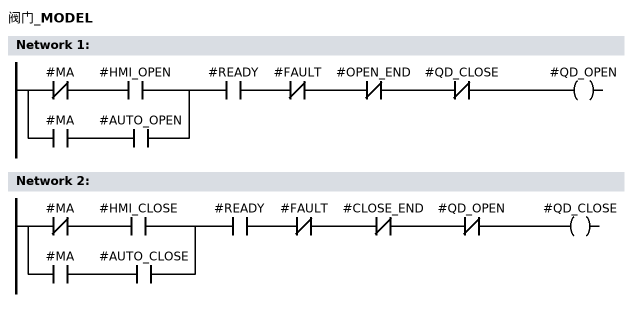
   RUNG wire#powerrail
      I_Contact( #MA )
      Contact( #HMI_OPEN )
      wire#w1
      Contact( #READY )
      I_Contact( #FAULT )
      I_Contact( #OPEN_END )
      I_Contact( #QD_CLOSE )
      Coil( #QD_OPEN )
   END_RUNG
   RUNG wire#powerrail
      Contact( #MA )
      Contact( #AUTO_OPEN )
   END_RUNG wire#w1
   // the same network as SCL:
   #QD_OPEN := ((NOT #MA AND #HMI_OPEN) OR (#MA AND #AUTO_OPEN)) AND #READY AND NOT #FAULT AND NOT #OPEN_END AND NOT #QD_CLOSE;
END_REGION

REGION Network 2
   RUNG wire#powerrail
      I_Contact( #MA )
      Contact( #HMI_CLOSE )
      wire#w1
      Contact( #READY )
      I_Contact( #FAULT )
      I_Contact( #CLOSE_END )
      I_Contact( #QD_OPEN )
      Coil( #QD_CLOSE )
   END_RUNG
   RUNG wire#powerrail
      Contact( #MA )
      Contact( #AUTO_CLOSE )
   END_RUNG wire#w1
   // the same network as SCL:
   #QD_CLOSE := ((NOT #MA AND #HMI_CLOSE) OR (#MA AND #AUTO_CLOSE)) AND #READY AND NOT #FAULT AND NOT #CLOSE_END AND NOT #QD_OPEN;
END_REGION
END_FUNCTION_BLOCK

FUNCTION_BLOCK "FB310_MOTOR_AUTO_ST_model"   // FB310, LAD
{ S7_Optimized_Access := 'FALSE' }
VERSION : 0.1
   VAR_INPUT
      LR_MOTOR : Bool;   // 水泵远程
      RUN_MOTOR : Bool;   // 水泵运行
      FAULT_MOTOR : Bool;   // 水泵故障
      LR_DF : Bool;   // 蝶阀远程
      FAULT_DF : Bool;   // 蝶阀故障
      CLOSE_END_DF : Bool;   // 蝶阀关到位
      HMI_AUTO : Bool;   // 画面选择自动
      HMI_MAN : Bool;   // 画面选择手动
      HMI_AUTO_ST : Bool;   // 画面自动启动
      HMI_AUTO_STP : Bool;   // 画面自动停止
      HMI_JT : Bool;   // 急停
      CX_AUTO_ST : Bool;   // 程序自动启动
      S : Bool;   // 0.5秒脉冲
      IN_T_ALARM : Time := T#15s;   // 报警时间
      IN_PT : Real;   // 压力
      IN_PT_QBYL : Real;   // 启泵压力
      IN_PT_KFYL : Real;   // 开阀压力,大于关泵压力
      IN_PT_GFYL : Real;   // 关阀压力
      IN_PT_DYYL : Real;   // 掉压压力
      IN_MOTRR_A : Real;   // 水泵电流
      IN_MOTOR_DYDL : Real;   // 掉压电流
      IN_TJFFK : Real;   // 调节阀反馈
   END_VAR
   VAR_IN_OUT
      OUT_AUTO : Bool;   // 自动模式
      AUTOING : Bool;   // 自动运行中
      OUT_FAULT : Bool;   // 自动模式故障
      OUT_ALARM : Bool;   // 报警输出
      OUT_PQF : Bool;   // 排气阀输出
      OUT_YSF : Bool;   // 引水阀输出
      OUT_MOTOR : Bool;   // 水泵输出
      OUT_DF_OPEN : Bool;   // 蝶阀开输出
      OUT_DF_CLOSE : Bool;   // 蝶阀关输出
      OUT_DF_CLOSE2 : Bool;   // 蝶阀关输出2
      OUT_QDXYT : Bool;   // 启动下一台输出
   END_VAR
   VAR
      T_ALARM : IEC_TIMER;
      T_MOTOR_RUN : IEC_TIMER;
      T_MOTOR_RUN2 : IEC_TIMER;
      T_MOTOR_RUN3 : IEC_TIMER;
      T_MOTOR_RUN4 : IEC_TIMER;
      P1 : Bool;
      P2 : Bool;
      P3 : Bool;
      P4 : Bool;
      P5 : Bool;
   END_VAR
   VAR_TEMP   // added for the SCL form of the ladder/FBD networks
      _w1 : Bool;
      _w2 : Bool;
   END_VAR
BEGIN

REGION Network 1: 自动模式
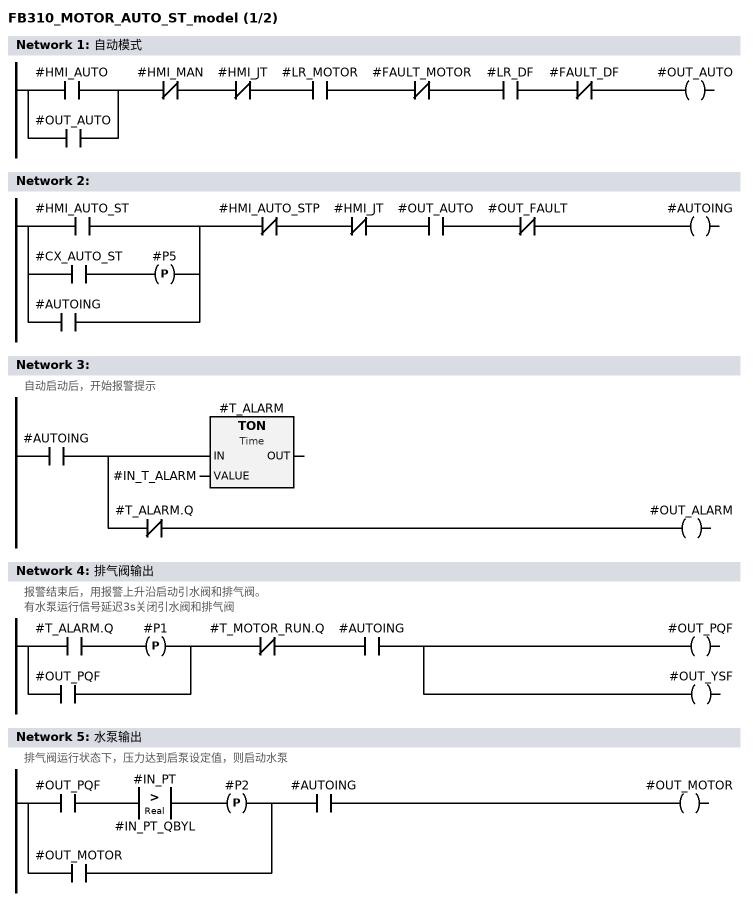
   RUNG wire#powerrail
      Contact( #HMI_AUTO )
      wire#w1
      I_Contact( #HMI_MAN )
      I_Contact( #HMI_JT )
      Contact( #LR_MOTOR )
      I_Contact( #FAULT_MOTOR )
      Contact( #LR_DF )
      I_Contact( #FAULT_DF )
      Coil( #OUT_AUTO )
   END_RUNG
   RUNG wire#powerrail
      Contact( #OUT_AUTO )
   END_RUNG wire#w1
   // the same network as SCL:
   #OUT_AUTO := (#HMI_AUTO OR #OUT_AUTO) AND NOT #HMI_MAN AND NOT #HMI_JT AND #LR_MOTOR AND NOT #FAULT_MOTOR AND #LR_DF AND NOT #FAULT_DF;
END_REGION

REGION Network 2
   RUNG wire#powerrail
      Contact( #HMI_AUTO_ST )
      wire#w1
      I_Contact( #HMI_AUTO_STP )
      I_Contact( #HMI_JT )
      Contact( #OUT_AUTO )
      I_Contact( #OUT_FAULT )
      Coil( #AUTOING )
   END_RUNG
   RUNG wire#powerrail
      Contact( #CX_AUTO_ST )
      P_Trig( #P5 )
   END_RUNG wire#w1
   RUNG wire#powerrail
      Contact( #AUTOING )
   END_RUNG wire#w1
   // the same network as SCL:
   #_w1 := #CX_AUTO_ST AND NOT #P5;   // rising edge
   #P5 := #CX_AUTO_ST;
   #AUTOING := (#HMI_AUTO_ST OR #_w1 OR #AUTOING) AND NOT #HMI_AUTO_STP AND NOT #HMI_JT AND #OUT_AUTO AND NOT #OUT_FAULT;
END_REGION

REGION Network 3
   // 自动启动后，开始报警提示
   #T_ALARM.TON(IN := #AUTOING, PT := #IN_T_ALARM);   // TON coil
   #OUT_ALARM := #AUTOING AND NOT #T_ALARM.Q;
END_REGION

REGION Network 4: 排气阀输出
   // 报警结束后，用报警上升沿启动引水阀和排气阀。
   // 有水泵运行信号延迟3s关闭引水阀和排气阀
   RUNG wire#powerrail
      Contact( #T_ALARM.Q )
      P_Trig( #P1 )
      wire#w1
      I_Contact( #T_MOTOR_RUN.Q )
      Contact( #AUTOING )
      wire#w2
      Coil( #OUT_PQF )
   END_RUNG
   RUNG wire#powerrail
      Contact( #OUT_PQF )
   END_RUNG wire#w1
   RUNG wire#w2
      Coil( #OUT_YSF )
   END_RUNG
   // the same network as SCL:
   #_w1 := #T_ALARM.Q AND NOT #P1;   // rising edge
   #P1 := #T_ALARM.Q;
   #OUT_PQF := (#_w1 OR #OUT_PQF) AND NOT #T_MOTOR_RUN.Q AND #AUTOING;
   #OUT_YSF := #OUT_PQF;
END_REGION

REGION Network 5: 水泵输出
   // 排气阀运行状态下，压力达到启泵设定值，则启动水泵
   RUNG wire#powerrail
      Contact( #OUT_PQF )
      { S7_Templates := "SrcType := Real" } GT_Contact(in1 := #IN_PT, in2 := #IN_PT_QBYL)
      P_Trig( #P2 )
      wire#w1
      Contact( #AUTOING )
      Coil( #OUT_MOTOR )
   END_RUNG
   RUNG wire#powerrail
      Contact( #OUT_MOTOR )
   END_RUNG wire#w1
   // the same network as SCL:
   #_w1 := #OUT_PQF AND (#IN_PT > #IN_PT_QBYL);
   #_w2 := #_w1 AND NOT #P2;   // rising edge
   #P2 := #_w1;
   #OUT_MOTOR := (#_w2 OR #OUT_MOTOR) AND #AUTOING;
END_REGION

REGION Network 6: 启动下一台输出
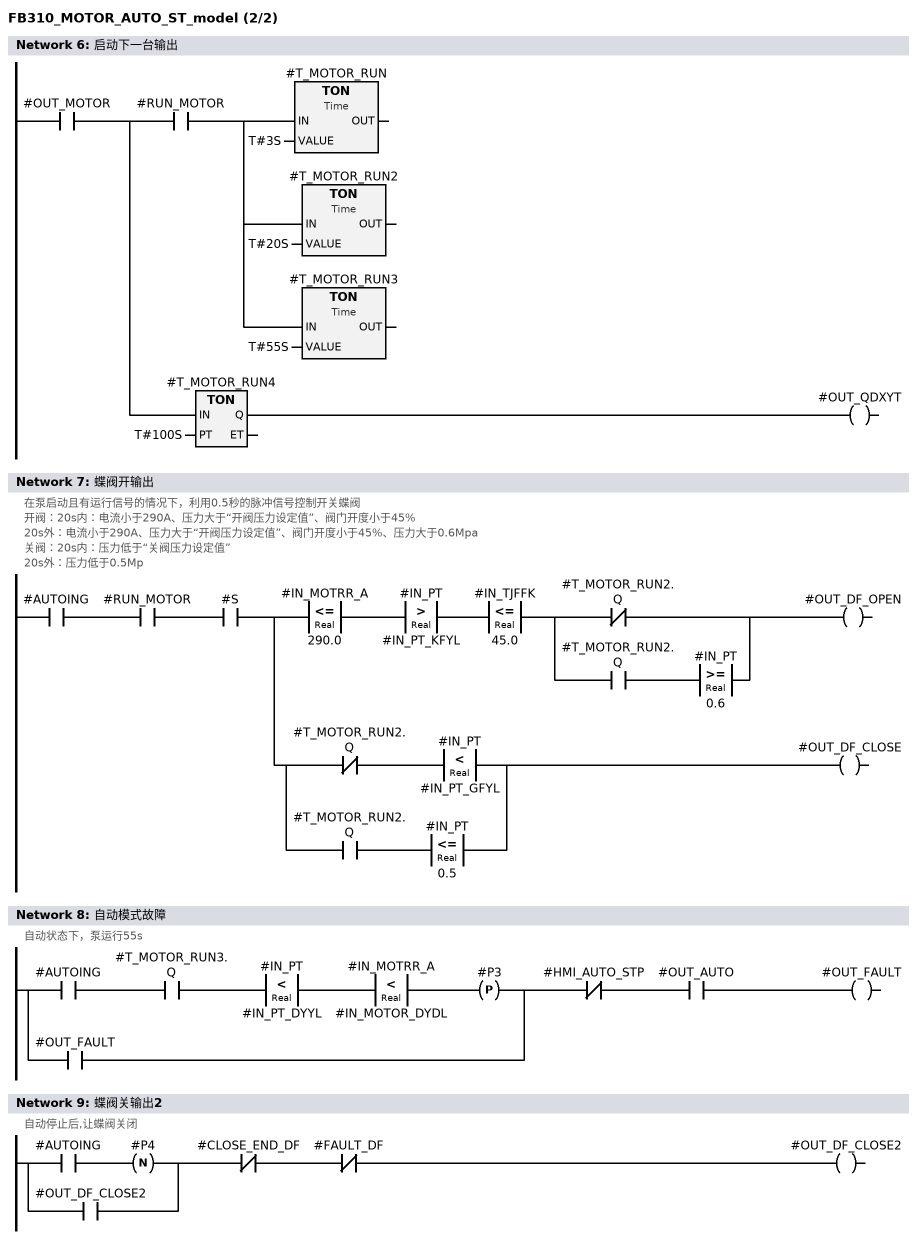
   #_w1 := #OUT_MOTOR AND #RUN_MOTOR;
   #T_MOTOR_RUN.TON(IN := #_w1, PT := T#3S);   // TON coil
   #T_MOTOR_RUN2.TON(IN := #_w1, PT := T#20S);   // TON coil
   #T_MOTOR_RUN3.TON(IN := #_w1, PT := T#55S);   // TON coil
   #T_MOTOR_RUN4.TON(IN := #OUT_MOTOR, PT := T#100S);
   #OUT_QDXYT := #T_MOTOR_RUN4.Q;
END_REGION

REGION Network 7: 蝶阀开输出
   // 在泵启动且有运行信号的情况下，利用0.5秒的脉冲信号控制开关蝶阀
   // 开阀：20s内：电流小于290A、压力大于“开阀压力设定值”、阀门开度小于45%
   //             20s外：电流小于290A、压力大于“开阀压力设定值”、阀门开度小于45%、压力大于0.6Mpa      
   // 关阀：20s内：压力低于“关阀压力设定值”
   //              20s外：压力低于0.5Mp
   RUNG wire#powerrail
      Contact( #AUTOING )
      Contact( #RUN_MOTOR )
      Contact( #S )
      wire#w1
      { S7_Templates := "SrcType := Real" } LE_Contact(in1 := #IN_MOTRR_A, in2 := 290.0)
      { S7_Templates := "SrcType := Real" } GT_Contact(in1 := #IN_PT, in2 := #IN_PT_KFYL)
      { S7_Templates := "SrcType := Real" } LE_Contact(in1 := #IN_TJFFK, in2 := 45.0)
      wire#w2
      I_Contact( #T_MOTOR_RUN2.Q )
      wire#w3
      Coil( #OUT_DF_OPEN )
   END_RUNG
   RUNG wire#w2
      Contact( #T_MOTOR_RUN2.Q )
      { S7_Templates := "SrcType := Real" } GE_Contact(in1 := #IN_PT, in2 := 0.6)
   END_RUNG wire#w3
   RUNG wire#w1
      I_Contact( #T_MOTOR_RUN2.Q )
      { S7_Templates := "SrcType := Real" } LT_Contact(in1 := #IN_PT, in2 := #IN_PT_GFYL)
      wire#w4
      Coil( #OUT_DF_CLOSE )
   END_RUNG
   RUNG wire#w1
      Contact( #T_MOTOR_RUN2.Q )
      { S7_Templates := "SrcType := Real" } LE_Contact(in1 := #IN_PT, in2 := 0.5)
   END_RUNG wire#w4
   // the same network as SCL:
   #_w1 := #AUTOING AND #RUN_MOTOR AND #S;
   #OUT_DF_OPEN := #_w1 AND (#IN_MOTRR_A <= 290.0) AND (#IN_PT > #IN_PT_KFYL) AND (#IN_TJFFK <= 45.0) AND (NOT #T_MOTOR_RUN2.Q OR (#T_MOTOR_RUN2.Q AND (#IN_PT >= 0.6)));
   #OUT_DF_CLOSE := #_w1 AND ((NOT #T_MOTOR_RUN2.Q AND (#IN_PT < #IN_PT_GFYL)) OR (#T_MOTOR_RUN2.Q AND (#IN_PT <= 0.5)));
END_REGION

REGION Network 8: 自动模式故障
   // 自动状态下，泵运行55s
   RUNG wire#powerrail
      Contact( #AUTOING )
      Contact( #T_MOTOR_RUN3.Q )
      { S7_Templates := "SrcType := Real" } LT_Contact(in1 := #IN_PT, in2 := #IN_PT_DYYL)
      { S7_Templates := "SrcType := Real" } LT_Contact(in1 := #IN_MOTRR_A, in2 := #IN_MOTOR_DYDL)
      P_Trig( #P3 )
      wire#w1
      I_Contact( #HMI_AUTO_STP )
      Contact( #OUT_AUTO )
      Coil( #OUT_FAULT )
   END_RUNG
   RUNG wire#powerrail
      Contact( #OUT_FAULT )
   END_RUNG wire#w1
   // the same network as SCL:
   #_w1 := #AUTOING AND #T_MOTOR_RUN3.Q AND (#IN_PT < #IN_PT_DYYL) AND (#IN_MOTRR_A < #IN_MOTOR_DYDL);
   #_w2 := #_w1 AND NOT #P3;   // rising edge
   #P3 := #_w1;
   #OUT_FAULT := (#_w2 OR #OUT_FAULT) AND NOT #HMI_AUTO_STP AND #OUT_AUTO;
END_REGION

REGION Network 9: 蝶阀关输出2
   // 自动停止后,让蝶阀关闭
   RUNG wire#powerrail
      Contact( #AUTOING )
      N_Trig( #P4 )
      wire#w1
      I_Contact( #CLOSE_END_DF )
      I_Contact( #FAULT_DF )
      Coil( #OUT_DF_CLOSE2 )
   END_RUNG
   RUNG wire#powerrail
      Contact( #OUT_DF_CLOSE2 )
   END_RUNG wire#w1
   // the same network as SCL:
   #_w1 := NOT #AUTOING AND #P4;   // falling edge
   #P4 := #AUTOING;
   #OUT_DF_CLOSE2 := (#_w1 OR #OUT_DF_CLOSE2) AND NOT #CLOSE_END_DF AND NOT #FAULT_DF;
END_REGION
END_FUNCTION_BLOCK

FUNCTION_BLOCK "引水排气块"   // FB320, LAD
{ S7_Optimized_Access := 'FALSE' }
VERSION : 0.1
// 阀门的手自动控制块
// 手动通过画面启停控制，带计时停止功能，且计时输出
// 自动通过自动控制信号控制，有则启动无则停止
   VAR_INPUT
      READY : Bool;
      HMI_OPEN : Bool;
      HMI_CLOSE : Bool;
      MA : Bool;
      AUTO : Bool;
      S : Bool;
      JT : Bool;
      "TIME" : Int := 15;
   END_VAR
   VAR_OUTPUT
      TIME_OUT : Int;   // 剩余时间
   END_VAR
   VAR_IN_OUT
      OUT : Bool;
   END_VAR
   VAR
      MAN_OUT : Bool;
      T_STOP : Bool;
      P1 : Bool;
      P2 : Bool;
      P3 : Bool;
      P4 : Bool;
      TIME_PV : Int;
   END_VAR
   VAR_TEMP   // added for the SCL form of the ladder/FBD networks
      _w1 : Bool;
      _w2 : Bool;
      _w3 : Bool;
   END_VAR
BEGIN

REGION Network 1
   // 手动输出，手动输出有计时
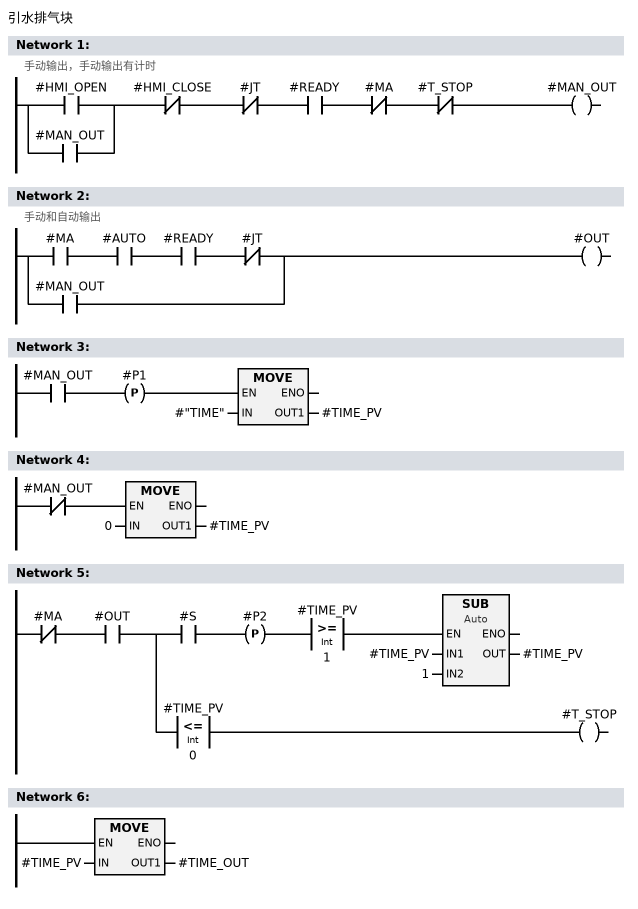
   RUNG wire#powerrail
      Contact( #HMI_OPEN )
      wire#w1
      I_Contact( #HMI_CLOSE )
      I_Contact( #JT )
      Contact( #READY )
      I_Contact( #MA )
      I_Contact( #T_STOP )
      Coil( #MAN_OUT )
   END_RUNG
   RUNG wire#powerrail
      Contact( #MAN_OUT )
   END_RUNG wire#w1
   // the same network as SCL:
   #MAN_OUT := (#HMI_OPEN OR #MAN_OUT) AND NOT #HMI_CLOSE AND NOT #JT AND #READY AND NOT #MA AND NOT #T_STOP;
END_REGION

REGION Network 2
   // 手动和自动输出
   RUNG wire#powerrail
      Contact( #MA )
      Contact( #AUTO )
      Contact( #READY )
      I_Contact( #JT )
      wire#w1
      Coil( #OUT )
   END_RUNG
   RUNG wire#powerrail
      Contact( #MAN_OUT )
   END_RUNG wire#w1
   // the same network as SCL:
   #OUT := (#MA AND #AUTO AND #READY AND NOT #JT) OR #MAN_OUT;
END_REGION

REGION Network 3
   RUNG wire#powerrail
      Contact( #MAN_OUT )
      P_Trig( #P1 )
      Move(in := #"TIME", out1 => #TIME_PV)
   END_RUNG
   // the same network as SCL:
   #_w1 := #MAN_OUT AND NOT #P1;   // rising edge
   #P1 := #MAN_OUT;
   IF #_w1 THEN #TIME_PV := #"TIME"; END_IF;
END_REGION

REGION Network 4
   RUNG wire#powerrail
      I_Contact( #MAN_OUT )
      Move(in := 0, out1 => #TIME_PV)
   END_RUNG
   // the same network as SCL:
   IF NOT #MAN_OUT THEN #TIME_PV := 0; END_IF;
END_REGION

REGION Network 5
   RUNG wire#powerrail
      I_Contact( #MA )
      Contact( #OUT )
      wire#w1
      Contact( #S )
      P_Trig( #P2 )
      { S7_Templates := "SrcType := Int" } GE_Contact(in1 := #TIME_PV, in2 := 1)
      Sub(in1 := #TIME_PV, in2 := 1, out => #TIME_PV)
   END_RUNG
   RUNG wire#w1
      { S7_Templates := "SrcType := Int" } LE_Contact(in1 := #TIME_PV, in2 := 0)
      Coil( #T_STOP )
   END_RUNG
   // the same network as SCL:
   #_w1 := NOT #MA AND #OUT;
   #_w2 := #_w1 AND #S;
   #_w3 := #_w2 AND NOT #P2;   // rising edge
   #P2 := #_w2;
   IF #_w3 AND (#TIME_PV >= 1) THEN #TIME_PV := #TIME_PV - 1; END_IF;
   #T_STOP := #_w1 AND (#TIME_PV <= 0);
END_REGION

REGION Network 6
   RUNG wire#powerrail
      Move(in := #TIME_PV, out1 => #TIME_OUT)
   END_RUNG
   // the same network as SCL:
   #TIME_OUT := #TIME_PV;
END_REGION
END_FUNCTION_BLOCK

FUNCTION_BLOCK "FB330_DATA_ALARM"   // FB330, LAD
{ S7_Optimized_Access := 'FALSE' }
VERSION : 0.1
// REAL的报警块
   VAR_INPUT
      PV : Real;   // 过程值
      PT : Real := 1.0;   // 系数
      HYS : Real;   // 回差值
      SV_AH : Real;   // 高报警设定值
      SV_WH : Real;   // 高警告设定值
      SV_WL : Real;   // 低警告设定值
      SV_AL : Real;   // 低报警设定值
      E_AH : Bool;   // 高报警使能
      E_WH : Bool;   // 高警告使能
      E_WL : Bool;   // 低警告使能
      E_AL : Bool;   // 低报警使能
   END_VAR
   VAR_OUTPUT
      QH_ALM : Bool;   // 高报警输出
      QH_WRN : Bool;   // 高警告输出
      QL_WRN : Bool;   // 低警告输出
      QL_ALM : Bool;   // 低报警输出
      OUT : Real;   // 输出
   END_VAR
   VAR
      SR1 : Bool;
      SR2 : Bool;
      SR3 : Bool;
      SR4 : Bool;
   END_VAR
   VAR_TEMP
      TEMP_AH : Real;
      TEMP_WH : Real;
      TEMP_AL : Real;
      TEMP_WL : Real;
      TEMP_OUT : Real;
   END_VAR
BEGIN

REGION Network 1
   // 系数转换
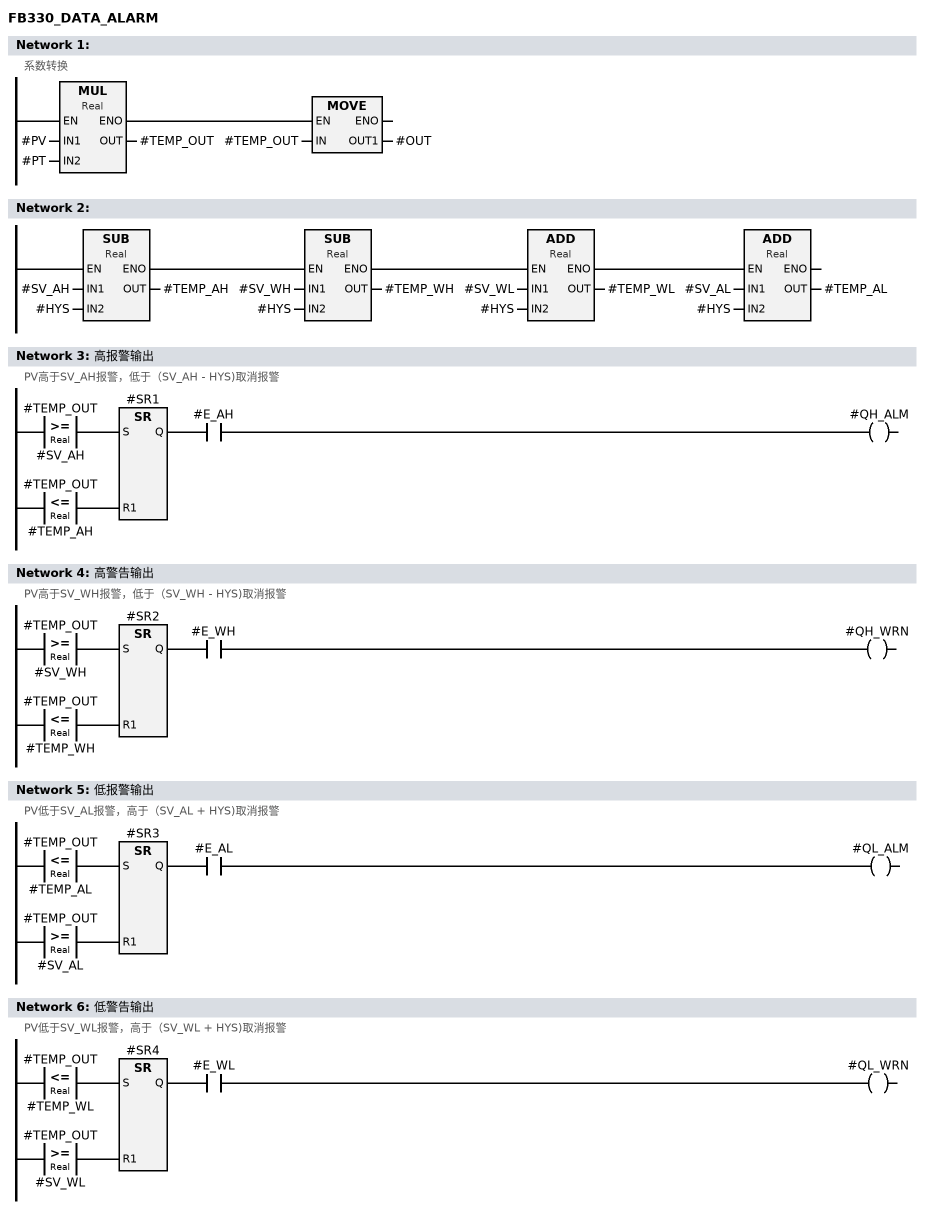
   RUNG wire#powerrail
      { S7_Templates := "SrcType := Real"; S7_GenerateENO := "TRUE" } Mul(in1 := #PV, in2 := #PT, out => #TEMP_OUT)
      { S7_GenerateENO := "TRUE" } Move(in := #TEMP_OUT, out1 => #OUT)
   END_RUNG
   // the same network as SCL:
   // ENO of a box is taken as its EN; it also drops when the box reports an error
   #TEMP_OUT := #PV * #PT;
   #OUT := #TEMP_OUT;
END_REGION

REGION Network 2
   RUNG wire#powerrail
      { S7_Templates := "SrcType := Real"; S7_GenerateENO := "TRUE" } Sub(in1 := #SV_AH, in2 := #HYS, out => #TEMP_AH)
      { S7_Templates := "SrcType := Real"; S7_GenerateENO := "TRUE" } Sub(in1 := #SV_WH, in2 := #HYS, out => #TEMP_WH)
      { S7_Templates := "SrcType := Real"; S7_GenerateENO := "TRUE" } Add(in1 := #SV_WL, in2 := #HYS, out => #TEMP_WL)
      { S7_Templates := "SrcType := Real"; S7_GenerateENO := "TRUE" } Add(in1 := #SV_AL, in2 := #HYS, out => #TEMP_AL)
   END_RUNG
   // the same network as SCL:
   // ENO of a box is taken as its EN; it also drops when the box reports an error
   #TEMP_AH := #SV_AH - #HYS;
   #TEMP_WH := #SV_WH - #HYS;
   #TEMP_WL := #SV_WL + #HYS;
   #TEMP_AL := #SV_AL + #HYS;
END_REGION

REGION Network 3: 高报警输出
   // PV高于SV_AH报警，低于（SV_AH - HYS)取消报警
   RUNG wire#powerrail
      { S7_Templates := "SrcType := Real" } GE_Contact(in1 := #TEMP_OUT, in2 := #SV_AH)
      S_SR(operand := #SR1, r1 := wire#w1)
      Contact( #E_AH )
      Coil( #QH_ALM )
   END_RUNG
   RUNG wire#powerrail
      { S7_Templates := "SrcType := Real" } LE_Contact(in1 := #TEMP_OUT, in2 := #TEMP_AH)
   END_RUNG wire#w1
   // the same network as SCL:
   IF #TEMP_OUT >= #SV_AH THEN
       #SR1 := TRUE;   // SR flip-flop
   END_IF;
   IF #TEMP_OUT <= #TEMP_AH THEN #SR1 := FALSE; END_IF;
   #QH_ALM := #SR1 AND #E_AH;
END_REGION

REGION Network 4: 高警告输出
   // PV高于SV_WH报警，低于（SV_WH - HYS)取消报警
   RUNG wire#powerrail
      { S7_Templates := "SrcType := Real" } GE_Contact(in1 := #TEMP_OUT, in2 := #SV_WH)
      S_SR(operand := #SR2, r1 := wire#w1)
      Contact( #E_WH )
      Coil( #QH_WRN )
   END_RUNG
   RUNG wire#powerrail
      { S7_Templates := "SrcType := Real" } LE_Contact(in1 := #TEMP_OUT, in2 := #TEMP_WH)
   END_RUNG wire#w1
   // the same network as SCL:
   IF #TEMP_OUT >= #SV_WH THEN
       #SR2 := TRUE;   // SR flip-flop
   END_IF;
   IF #TEMP_OUT <= #TEMP_WH THEN #SR2 := FALSE; END_IF;
   #QH_WRN := #SR2 AND #E_WH;
END_REGION

REGION Network 5: 低报警输出
   // PV低于SV_AL报警，高于（SV_AL + HYS)取消报警
   RUNG wire#powerrail
      { S7_Templates := "SrcType := Real" } LE_Contact(in1 := #TEMP_OUT, in2 := #TEMP_AL)
      S_SR(operand := #SR3, r1 := wire#w1)
      Contact( #E_AL )
      Coil( #QL_ALM )
   END_RUNG
   RUNG wire#powerrail
      { S7_Templates := "SrcType := Real" } GE_Contact(in1 := #TEMP_OUT, in2 := #SV_AL)
   END_RUNG wire#w1
   // the same network as SCL:
   IF #TEMP_OUT <= #TEMP_AL THEN
       #SR3 := TRUE;   // SR flip-flop
   END_IF;
   IF #TEMP_OUT >= #SV_AL THEN #SR3 := FALSE; END_IF;
   #QL_ALM := #SR3 AND #E_AL;
END_REGION

REGION Network 6: 低警告输出
   // PV低于SV_WL报警，高于（SV_WL + HYS)取消报警
   RUNG wire#powerrail
      { S7_Templates := "SrcType := Real" } LE_Contact(in1 := #TEMP_OUT, in2 := #TEMP_WL)
      S_SR(operand := #SR4, r1 := wire#w1)
      Contact( #E_WL )
      Coil( #QL_WRN )
   END_RUNG
   RUNG wire#powerrail
      { S7_Templates := "SrcType := Real" } GE_Contact(in1 := #TEMP_OUT, in2 := #SV_WL)
   END_RUNG wire#w1
   // the same network as SCL:
   IF #TEMP_OUT <= #TEMP_WL THEN
       #SR4 := TRUE;   // SR flip-flop
   END_IF;
   IF #TEMP_OUT >= #SV_WL THEN #SR4 := FALSE; END_IF;
   #QL_WRN := #SR4 AND #E_WL;
END_REGION
END_FUNCTION_BLOCK

FUNCTION_BLOCK "流量累计块2"   // FB331, LAD
{ S7_Optimized_Access := 'FALSE' }
VERSION : 0.1
// 模拟量的累计，每100ms加一次数值。
// 数值精确到小数位后两位。
// 累计上线555.5
   VAR_INPUT
      FIT : Real;
      CLEAR1 : Bool;
      CLEAR2 : Bool;
      CLEAR3 : Bool;
   END_VAR
   VAR_OUTPUT
      OUT1 : Real;
      OUT2 : Real;
      OUT3 : Real;
   END_VAR
   VAR
      STATIC1 : Real;
      TEMP_STATIC : DInt;
      FQIT1 : DInt;
      FQIT2 : DInt;
      FQIT3 : DInt;
      FQIT1_2 : Real;
      FQIT2_2 : Real;
      FQIT3_2 : Real;
   END_VAR
BEGIN

REGION Network 1
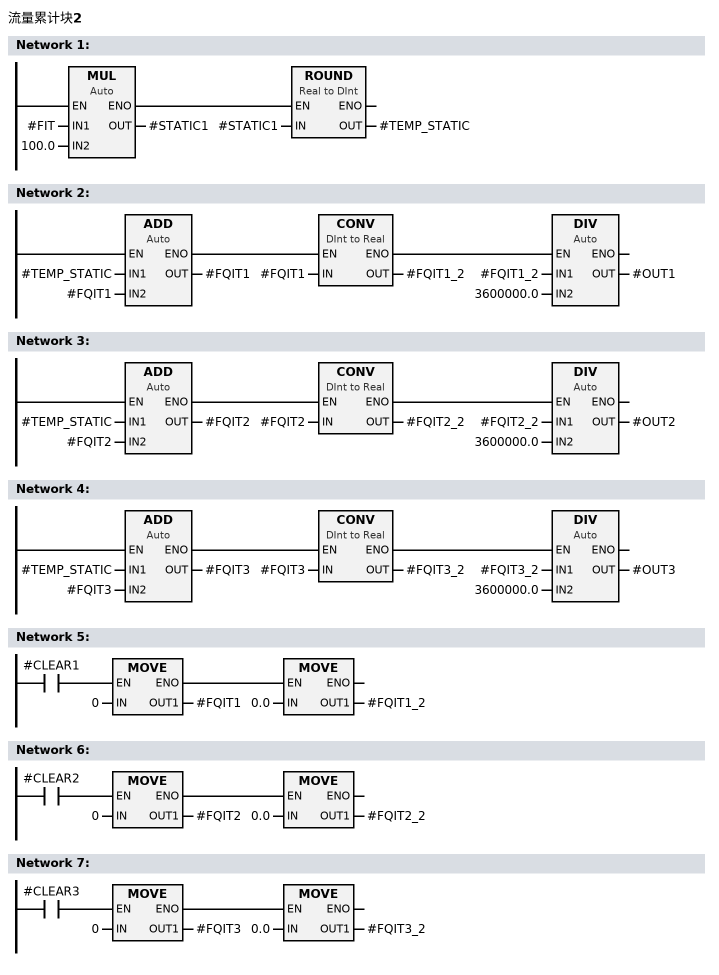
   RUNG wire#powerrail
      Mul(in1 := #FIT, in2 := 100.0, out => #STATIC1)
      { S7_Templates := "[SrcType := Real, DestType := DInt]" } Round(in := #STATIC1, out => #TEMP_STATIC)
   END_RUNG
   // the same network as SCL:
   #STATIC1 := #FIT * 100.0;
   #TEMP_STATIC := ROUND(#STATIC1);
END_REGION

REGION Network 2
   RUNG wire#powerrail
      Add(in1 := #TEMP_STATIC, in2 := #FQIT1, out => #FQIT1)
      { S7_Templates := "[SrcType := DInt, DestType := Real]" } Convert(in := #FQIT1, out => #FQIT1_2)
      Div(in1 := #FQIT1_2, in2 := 3600000.0, out => #OUT1)
   END_RUNG
   // the same network as SCL:
   #FQIT1 := #TEMP_STATIC + #FQIT1;
   #FQIT1_2 := DINT_TO_REAL(#FQIT1);
   #OUT1 := #FQIT1_2 / 3600000.0;
END_REGION

REGION Network 3
   RUNG wire#powerrail
      Add(in1 := #TEMP_STATIC, in2 := #FQIT2, out => #FQIT2)
      { S7_Templates := "[SrcType := DInt, DestType := Real]" } Convert(in := #FQIT2, out => #FQIT2_2)
      Div(in1 := #FQIT2_2, in2 := 3600000.0, out => #OUT2)
   END_RUNG
   // the same network as SCL:
   #FQIT2 := #TEMP_STATIC + #FQIT2;
   #FQIT2_2 := DINT_TO_REAL(#FQIT2);
   #OUT2 := #FQIT2_2 / 3600000.0;
END_REGION

REGION Network 4
   RUNG wire#powerrail
      Add(in1 := #TEMP_STATIC, in2 := #FQIT3, out => #FQIT3)
      { S7_Templates := "[SrcType := DInt, DestType := Real]" } Convert(in := #FQIT3, out => #FQIT3_2)
      Div(in1 := #FQIT3_2, in2 := 3600000.0, out => #OUT3)
   END_RUNG
   // the same network as SCL:
   #FQIT3 := #TEMP_STATIC + #FQIT3;
   #FQIT3_2 := DINT_TO_REAL(#FQIT3);
   #OUT3 := #FQIT3_2 / 3600000.0;
END_REGION

REGION Network 5
   RUNG wire#powerrail
      Contact( #CLEAR1 )
      Move(in := 0, out1 => #FQIT1)
      Move(in := 0.0, out1 => #FQIT1_2)
   END_RUNG
   // the same network as SCL:
   IF #CLEAR1 THEN
       #FQIT1 := 0;
       #FQIT1_2 := 0.0;
   END_IF;
END_REGION

REGION Network 6
   RUNG wire#powerrail
      Contact( #CLEAR2 )
      Move(in := 0, out1 => #FQIT2)
      Move(in := 0.0, out1 => #FQIT2_2)
   END_RUNG
   // the same network as SCL:
   IF #CLEAR2 THEN
       #FQIT2 := 0;
       #FQIT2_2 := 0.0;
   END_IF;
END_REGION

REGION Network 7
   RUNG wire#powerrail
      Contact( #CLEAR3 )
      Move(in := 0, out1 => #FQIT3)
      Move(in := 0.0, out1 => #FQIT3_2)
   END_RUNG
   // the same network as SCL:
   IF #CLEAR3 THEN
       #FQIT3 := 0;
       #FQIT3_2 := 0.0;
   END_IF;
END_REGION
END_FUNCTION_BLOCK

FUNCTION "FC1_模拟量输入" : Void   // FC1, LAD
{ S7_Optimized_Access := 'TRUE' }
VERSION : 0.1
   VAR_TEMP
      temp : Word;
   END_VAR
BEGIN

REGION Network 1
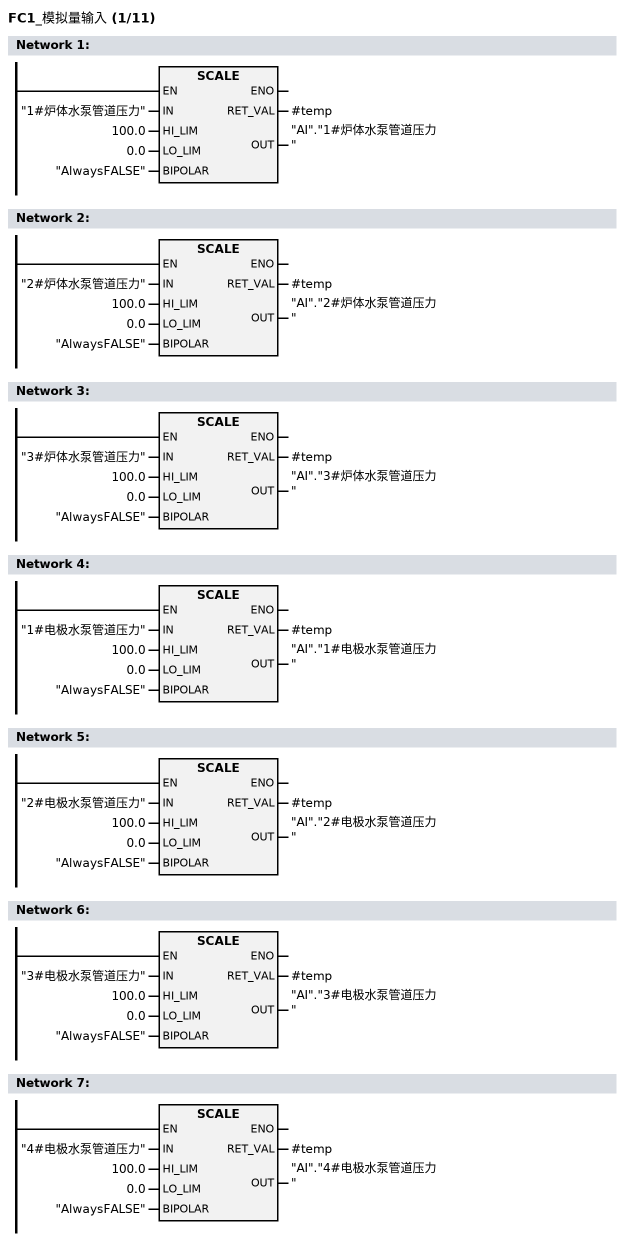
   #temp := SCALE(IN := "1#炉体水泵管道压力",
                  HI_LIM := 100.0,
                  LO_LIM := 0.0,
                  BIPOLAR := "AlwaysFALSE",
                  OUT => "AI"."1#炉体水泵管道压力");
END_REGION

REGION Network 2
   #temp := SCALE(IN := "2#炉体水泵管道压力",
                  HI_LIM := 100.0,
                  LO_LIM := 0.0,
                  BIPOLAR := "AlwaysFALSE",
                  OUT => "AI"."2#炉体水泵管道压力");
END_REGION

REGION Network 3
   #temp := SCALE(IN := "3#炉体水泵管道压力",
                  HI_LIM := 100.0,
                  LO_LIM := 0.0,
                  BIPOLAR := "AlwaysFALSE",
                  OUT => "AI"."3#炉体水泵管道压力");
END_REGION

REGION Network 4
   #temp := SCALE(IN := "1#电极水泵管道压力",
                  HI_LIM := 100.0,
                  LO_LIM := 0.0,
                  BIPOLAR := "AlwaysFALSE",
                  OUT => "AI"."1#电极水泵管道压力");
END_REGION

REGION Network 5
   #temp := SCALE(IN := "2#电极水泵管道压力",
                  HI_LIM := 100.0,
                  LO_LIM := 0.0,
                  BIPOLAR := "AlwaysFALSE",
                  OUT => "AI"."2#电极水泵管道压力");
END_REGION

REGION Network 6
   #temp := SCALE(IN := "3#电极水泵管道压力",
                  HI_LIM := 100.0,
                  LO_LIM := 0.0,
                  BIPOLAR := "AlwaysFALSE",
                  OUT => "AI"."3#电极水泵管道压力");
END_REGION

REGION Network 7
   #temp := SCALE(IN := "4#电极水泵管道压力",
                  HI_LIM := 100.0,
                  LO_LIM := 0.0,
                  BIPOLAR := "AlwaysFALSE",
                  OUT => "AI"."4#电极水泵管道压力");
END_REGION

REGION Network 8
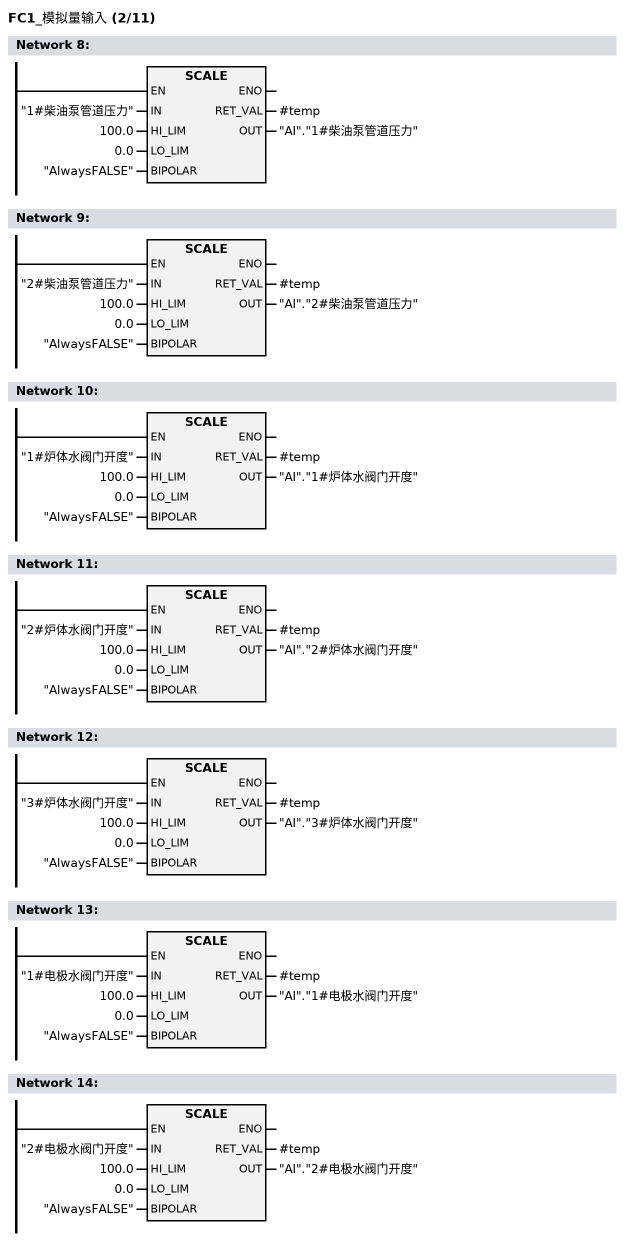
   #temp := SCALE(IN := "1#柴油泵管道压力",
                  HI_LIM := 100.0,
                  LO_LIM := 0.0,
                  BIPOLAR := "AlwaysFALSE",
                  OUT => "AI"."1#柴油泵管道压力");
END_REGION

REGION Network 9
   #temp := SCALE(IN := "2#柴油泵管道压力",
                  HI_LIM := 100.0,
                  LO_LIM := 0.0,
                  BIPOLAR := "AlwaysFALSE",
                  OUT => "AI"."2#柴油泵管道压力");
END_REGION

REGION Network 10
   #temp := SCALE(IN := "1#炉体水阀门开度",
                  HI_LIM := 100.0,
                  LO_LIM := 0.0,
                  BIPOLAR := "AlwaysFALSE",
                  OUT => "AI"."1#炉体水阀门开度");
END_REGION

REGION Network 11
   #temp := SCALE(IN := "2#炉体水阀门开度",
                  HI_LIM := 100.0,
                  LO_LIM := 0.0,
                  BIPOLAR := "AlwaysFALSE",
                  OUT => "AI"."2#炉体水阀门开度");
END_REGION

REGION Network 12
   #temp := SCALE(IN := "3#炉体水阀门开度",
                  HI_LIM := 100.0,
                  LO_LIM := 0.0,
                  BIPOLAR := "AlwaysFALSE",
                  OUT => "AI"."3#炉体水阀门开度");
END_REGION

REGION Network 13
   #temp := SCALE(IN := "1#电极水阀门开度",
                  HI_LIM := 100.0,
                  LO_LIM := 0.0,
                  BIPOLAR := "AlwaysFALSE",
                  OUT => "AI"."1#电极水阀门开度");
END_REGION

REGION Network 14
   #temp := SCALE(IN := "2#电极水阀门开度",
                  HI_LIM := 100.0,
                  LO_LIM := 0.0,
                  BIPOLAR := "AlwaysFALSE",
                  OUT => "AI"."2#电极水阀门开度");
END_REGION

REGION Network 15
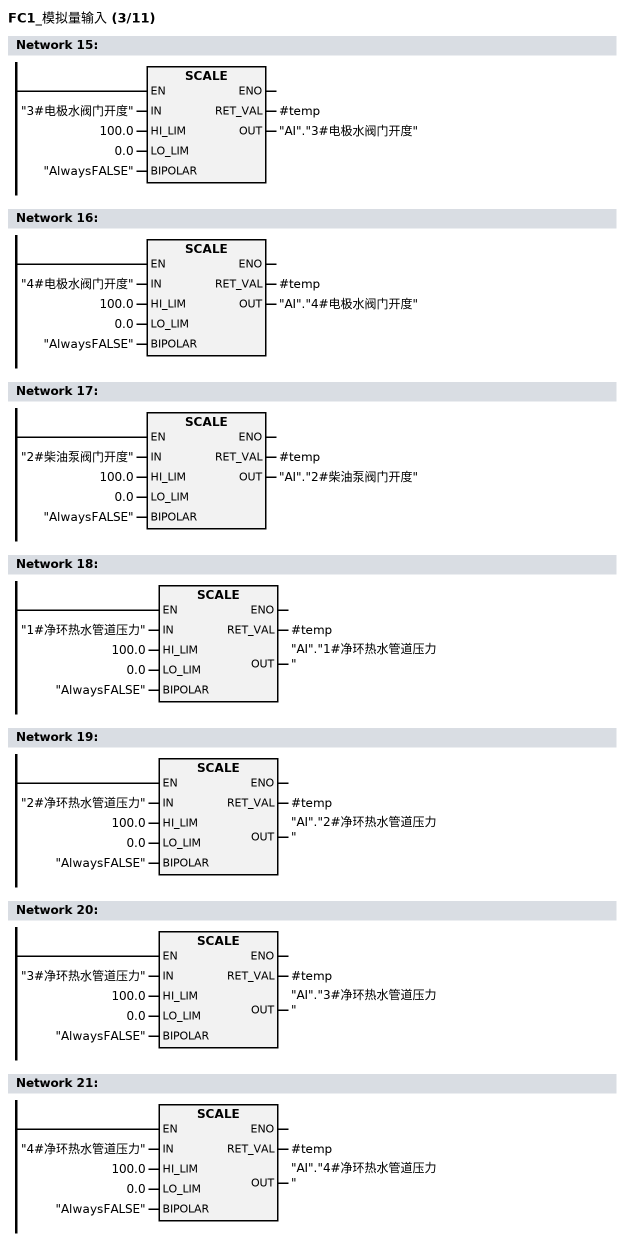
   #temp := SCALE(IN := "3#电极水阀门开度",
                  HI_LIM := 100.0,
                  LO_LIM := 0.0,
                  BIPOLAR := "AlwaysFALSE",
                  OUT => "AI"."3#电极水阀门开度");
END_REGION

REGION Network 16
   #temp := SCALE(IN := "4#电极水阀门开度",
                  HI_LIM := 100.0,
                  LO_LIM := 0.0,
                  BIPOLAR := "AlwaysFALSE",
                  OUT => "AI"."4#电极水阀门开度");
END_REGION

REGION Network 17
   #temp := SCALE(IN := "2#柴油泵阀门开度",
                  HI_LIM := 100.0,
                  LO_LIM := 0.0,
                  BIPOLAR := "AlwaysFALSE",
                  OUT => "AI"."2#柴油泵阀门开度");
END_REGION

REGION Network 18
   #temp := SCALE(IN := "1#净环热水管道压力",
                  HI_LIM := 100.0,
                  LO_LIM := 0.0,
                  BIPOLAR := "AlwaysFALSE",
                  OUT => "AI"."1#净环热水管道压力");
END_REGION

REGION Network 19
   #temp := SCALE(IN := "2#净环热水管道压力",
                  HI_LIM := 100.0,
                  LO_LIM := 0.0,
                  BIPOLAR := "AlwaysFALSE",
                  OUT => "AI"."2#净环热水管道压力");
END_REGION

REGION Network 20
   #temp := SCALE(IN := "3#净环热水管道压力",
                  HI_LIM := 100.0,
                  LO_LIM := 0.0,
                  BIPOLAR := "AlwaysFALSE",
                  OUT => "AI"."3#净环热水管道压力");
END_REGION

REGION Network 21
   #temp := SCALE(IN := "4#净环热水管道压力",
                  HI_LIM := 100.0,
                  LO_LIM := 0.0,
                  BIPOLAR := "AlwaysFALSE",
                  OUT => "AI"."4#净环热水管道压力");
END_REGION

REGION Network 22
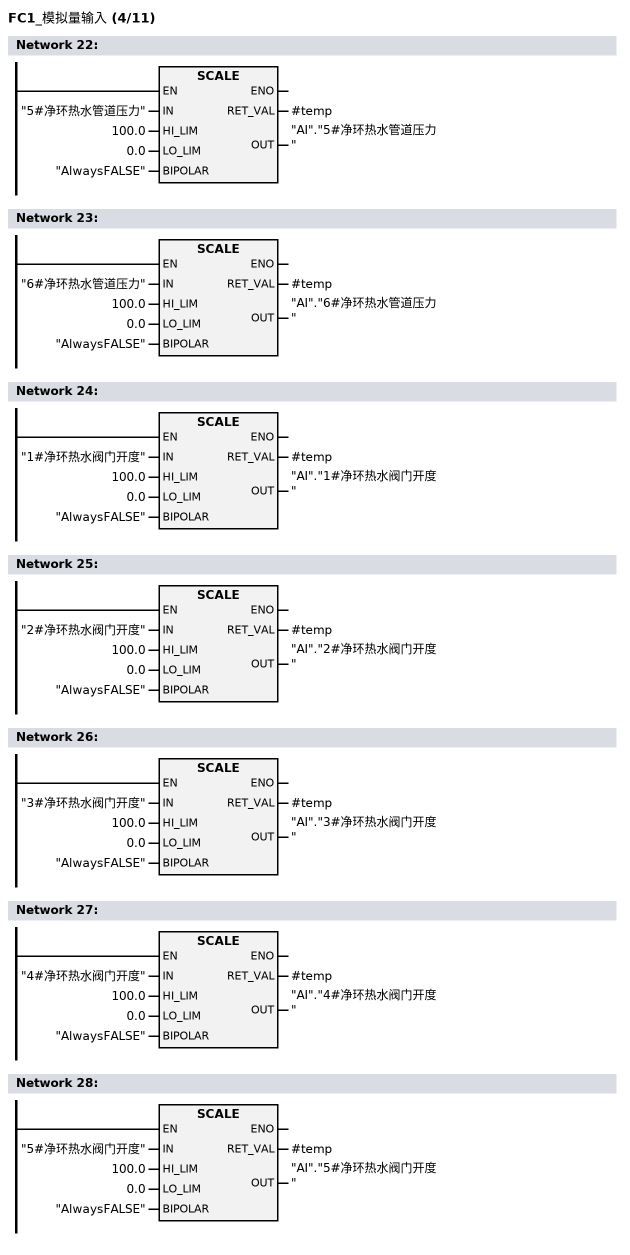
   #temp := SCALE(IN := "5#净环热水管道压力",
                  HI_LIM := 100.0,
                  LO_LIM := 0.0,
                  BIPOLAR := "AlwaysFALSE",
                  OUT => "AI"."5#净环热水管道压力");
END_REGION

REGION Network 23
   #temp := SCALE(IN := "6#净环热水管道压力",
                  HI_LIM := 100.0,
                  LO_LIM := 0.0,
                  BIPOLAR := "AlwaysFALSE",
                  OUT => "AI"."6#净环热水管道压力");
END_REGION

REGION Network 24
   #temp := SCALE(IN := "1#净环热水阀门开度",
                  HI_LIM := 100.0,
                  LO_LIM := 0.0,
                  BIPOLAR := "AlwaysFALSE",
                  OUT => "AI"."1#净环热水阀门开度");
END_REGION

REGION Network 25
   #temp := SCALE(IN := "2#净环热水阀门开度",
                  HI_LIM := 100.0,
                  LO_LIM := 0.0,
                  BIPOLAR := "AlwaysFALSE",
                  OUT => "AI"."2#净环热水阀门开度");
END_REGION

REGION Network 26
   #temp := SCALE(IN := "3#净环热水阀门开度",
                  HI_LIM := 100.0,
                  LO_LIM := 0.0,
                  BIPOLAR := "AlwaysFALSE",
                  OUT => "AI"."3#净环热水阀门开度");
END_REGION

REGION Network 27
   #temp := SCALE(IN := "4#净环热水阀门开度",
                  HI_LIM := 100.0,
                  LO_LIM := 0.0,
                  BIPOLAR := "AlwaysFALSE",
                  OUT => "AI"."4#净环热水阀门开度");
END_REGION
